   X1_BLTS_PROCS : ALIAS FOR I[3].0;
   XFER1A_BLTS_PRO : ALIAS FOR I[3].6;
   Z200 : MAC_Zone_ML := (ST_xManualModeConditionOK := 1, ST_xZoneError := 1, tmON_480Vca.ACC := 10, tmON_480Vca.EN := 1, tmON_480Vca.DN := 1);
   Z200_ALM : MAC_Zone_ML_ALM := (rgxEmergency[0] := 1, rgxStoppingFault[0] := 63, rgxWarning[0] := 7);
        .rgxEmergency[0].0   // MCC1201.A34KE1.Main Emergency ON
        .rgxStoppingFault[0].0   // Z200.MCC1201.24Vdc Voltage Fault
        .rgxEmergency[0].1   // MCC1201.A33SB1.Main Emergency localization (MCC1201 cabinet)
        .rgxEmergency[0].2   // M203S.A34SB1.Main Emergency localization (operator side)
        .rgxEmergency[0].3   // M203S.A34SB2.Main Emergency localization (far side)
        .rgxStoppingFault[0].1   // Z200.MCC1201.A18QF31/32/33/34.Power supply 24Vdc Fault
        .rgxStoppingFault[0].2   // Z200.MCC1201.A18QF41/42/43/44.Power supply 24Vdc Fault
        .rgxStoppingFault[0].3   // Z200.MCC1201.A19QF11/12/13/14.Power supply 24Vdc Fault
        .rgxStoppingFault[0].4   // Z200.MCC1201.A19QF21/22/23/24.Power supply 24Vdc Fault
        .rgxFault[0].0   // Z200.MCC1201.A155SW1.Ethernet Switch Fault
        .rgxWarning[0].0   // Z200.MCC1201.A11QF1.Power failure 120V Auxiliary
        .rgxWarning[0].1   // Z200.MCC1201.A11QF3.Power failure 120V Auxiliary
        .rgxWarning[0].2   // Z200.MCC1201.A16QF1.Protection power supply conditioner
        .rgxStoppingFault[0].5   // Z200.MCC1201.A18GS1.24Vdc Power Supply Fault
   Z200_HMR : MAC_Zone_ML_HMR := (xZoneAlarm := 1, dZoneState := 1024, dCabinetState := 2, dCleaningState := 2, dManualSpeed_mm_min := 1270);
   Z200_HMW : MAC_Zone_ML_HMW;
   Z200_UPS : ZONE_UPS := (ST_xZoneError := 1, ST_xSelectionManualMode := 1, ST_xConditionOKManualMode := 1, ST_xManualModeAccepted := 1, ST_xZoneEmergency := 1, INPUT_xPowerFailurePLCA := 1, INPUT_xPowerFailurePLCB := 1, AUX_tmOFF_ResetAlarm.PRE := 1000, AUX_tmOFF_ResetAlarm.ACC := 1000, AUX_tmON_24Vdc.PRE := 5000, AUX_tmON_EmergencyOK.PRE := 5000, AUX_tmON_Clutch1feedback.PRE := 1000, AUX_tmON_Clutch2feedback.PRE := 1000); {access None}
   Z200_UPS_ALM : ZONE_UPS_ALM := (rgxEmergency[0] := 1); {access Read Only}
        .rgxEmergency[0].0   // MCC1201.A33KE1.UPS Emergency ON
        .rgxEmergency[0].1   // M203S.A33SB2.UPS Emergency localization (operator side)
        .rgxEmergency[0].2   // M203S.A33SB3.UPS Emergency localization (far side)
        .rgxEmergency[0].3   // M225S.A33SB4.UPS Emergency localization (operator side CS4425)
        .rgxEmergency[0].4   // M225S.A33SB5.UPS Emergency localization (operator side CS4425)
   Z200_UPS_HMR : ZONE_UPS_HMR := (dZoneMode := 1, xZoneAlarm := 1, dZoneState := 1024); {access Read Only}
   Z200_UPS_HMW : ZONE_UPS_HMW;
   Z_ONS_BIT : BOOL[32];   // Temporary Boolean tag created during conversion
END_VAR

PROGRAM _18_STI   (* main routine _18_STI *)

ROUTINE _18_STI   (* ladder *)
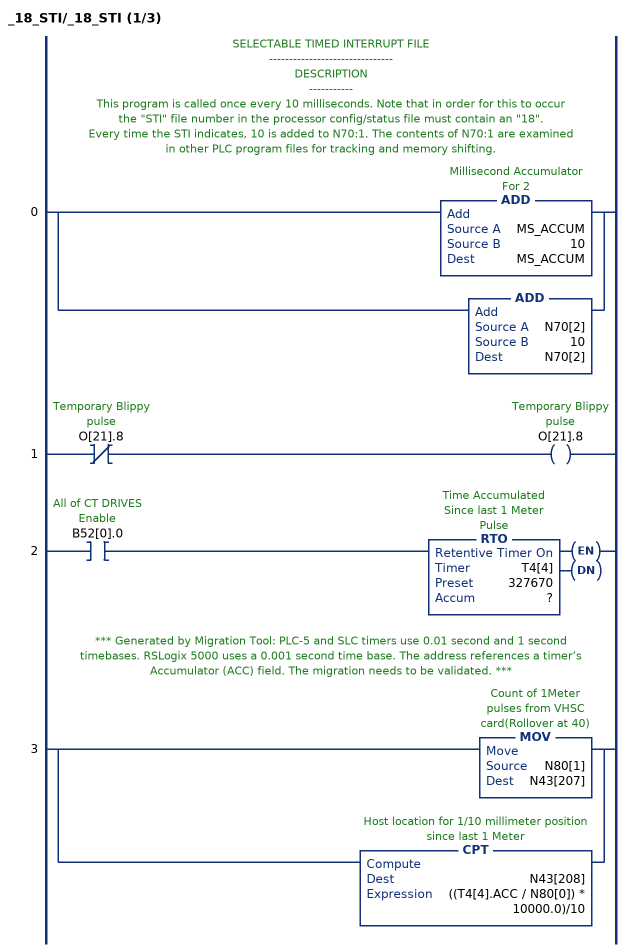
   // SELECTABLE TIMED INTERRUPT FILE
   // -------------------------------
   // DESCRIPTION
   // -----------
   // This program is called once every 10 milliseconds. Note that in order for this to occur
   // the "STI" file number in the processor config/status file must contain an "18".
   // Every time the STI indicates, 10 is added to N70:1. The contents of N70:1 are examined
   // in other PLC program files for tracking and memory shifting.
   0: [ADD(MS_ACCUM,10,MS_ACCUM) ,ADD(N70[2],10,N70[2]) ];
   1: XIO(O[21].8)OTE(O[21].8);
   2: XIC(B52[0].0)RTO(T4[4],?,?);
   // *** Generated by Migration Tool: PLC-5 and SLC timers use 0.01 second and 1 second timebases. RSLogix 5000 uses a 0.001 second time base. The address references a timer’s Accumulator (ACC) field. The migration needs to be validated. ***
   3: [MOV(N80[1],N43[207]) ,CPT(N43[208],((T4[4].ACC / N80[0]) * 10000.0)/10) ];
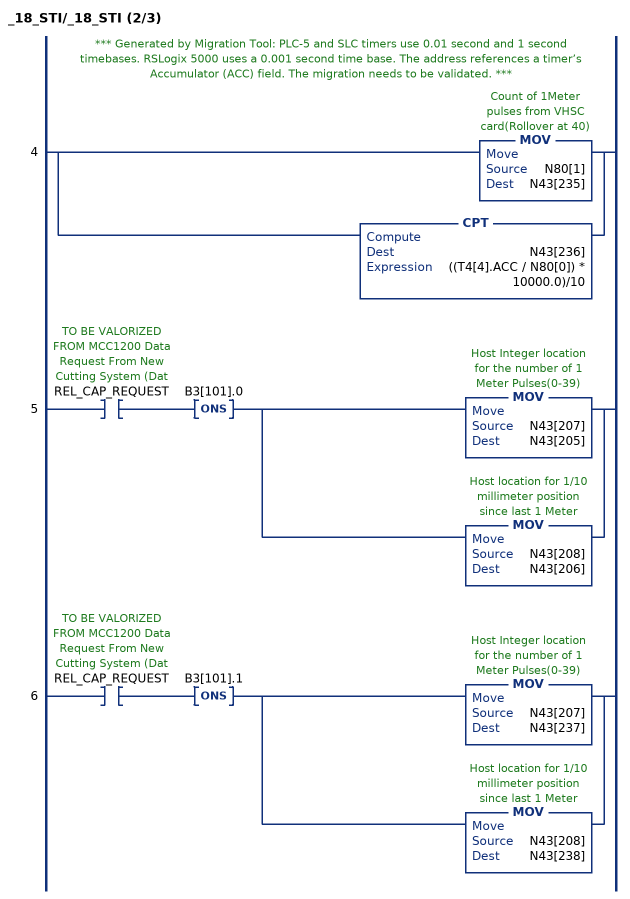
   // *** Generated by Migration Tool: PLC-5 and SLC timers use 0.01 second and 1 second timebases. RSLogix 5000 uses a 0.001 second time base. The address references a timer’s Accumulator (ACC) field. The migration needs to be validated. ***
   4: [MOV(N80[1],N43[235]) ,CPT(N43[236],((T4[4].ACC / N80[0]) * 10000.0)/10) ];
   5: XIC(REL_CAP_REQUEST)ONS(B3[101].0)[MOV(N43[207],N43[205]) ,MOV(N43[208],N43[206]) ];
   6: XIC(REL_CAP_REQUEST)ONS(B3[101].1)[MOV(N43[207],N43[237]) ,MOV(N43[208],N43[238]) ];
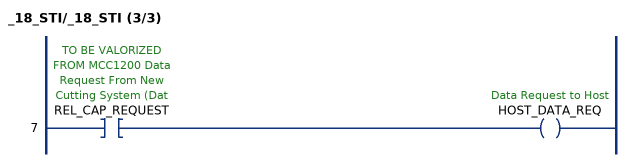
   7: XIC(REL_CAP_REQUEST)OTE(HOST_DATA_REQ);
END_ROUTINE
END_PROGRAM

PROGRAM CommandLogic   (* main routine Main *)
VAR
   TMP_rDummy : REAL;
   TMP_rTarget : REAL;
   TMP_xDummy : BOOL;
   WASHER_ALARM_HORN_RESET : BOOL;
END_VAR

ROUTINE M202_Conveyor_Motion_Output   (* ladder *)
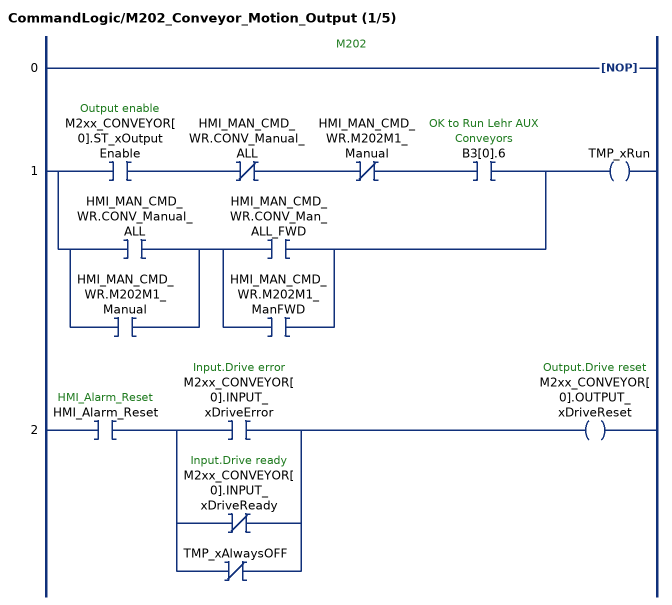
   // M202
   0: NOP();
   1: [XIC(M2xx_CONVEYOR[0].ST_xOutputEnable) XIO(HMI_MAN_CMD_WR.CONV_Manual_ALL) XIO(HMI_MAN_CMD_WR.M202M1_Manual) XIC(B3[0].6) ,[XIC(HMI_MAN_CMD_WR.CONV_Manual_ALL) ,XIC(HMI_MAN_CMD_WR.M202M1_Manual) ] [XIC(HMI_MAN_CMD_WR.CONV_Man_ALL_FWD) ,XIC(HMI_MAN_CMD_WR.M202M1_ManFWD) ] ]OTE(TMP_xRun);
   2: XIC(HMI_Alarm_Reset)[XIC(M2xx_CONVEYOR[0].INPUT_xDriveError) ,XIO(M2xx_CONVEYOR[0].INPUT_xDriveReady) ,XIO(TMP_xAlwaysOFF) ]OTE(M2xx_CONVEYOR[0].OUTPUT_xDriveReset);
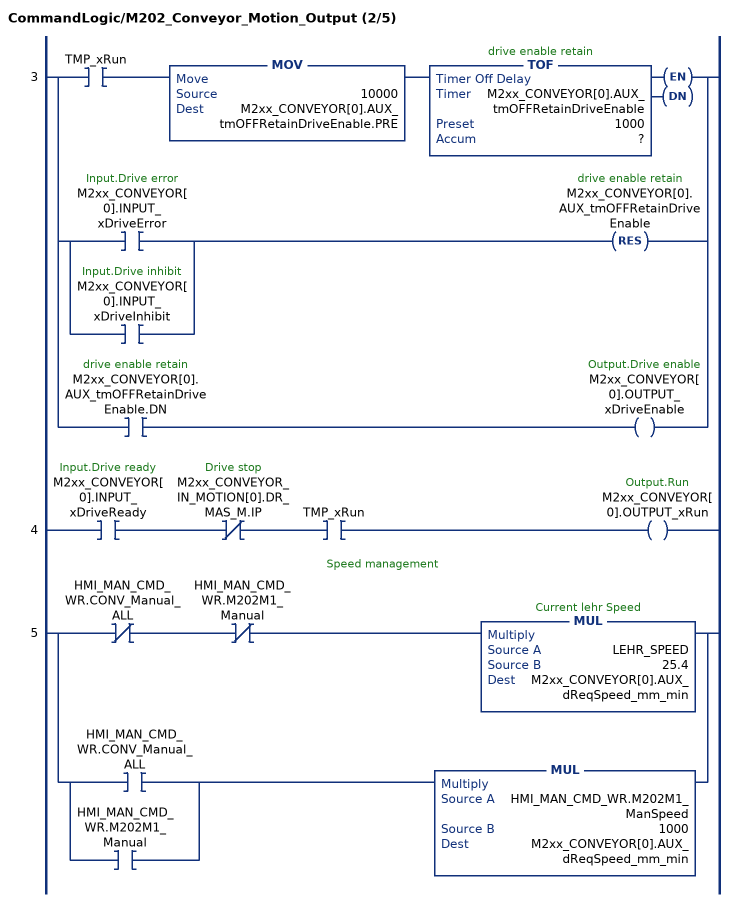
   3: [XIC(TMP_xRun) MOV(10000,M2xx_CONVEYOR[0].AUX_tmOFFRetainDriveEnable.PRE) TOF(M2xx_CONVEYOR[0].AUX_tmOFFRetainDriveEnable,?,?) ,[XIC(M2xx_CONVEYOR[0].INPUT_xDriveError) ,XIC(M2xx_CONVEYOR[0].INPUT_xDriveInhibit) ] RES(M2xx_CONVEYOR[0].AUX_tmOFFRetainDriveEnable) ,XIC(M2xx_CONVEYOR[0].AUX_tmOFFRetainDriveEnable.DN) OTE(M2xx_CONVEYOR[0].OUTPUT_xDriveEnable) ];
   4: XIC(M2xx_CONVEYOR[0].INPUT_xDriveReady)XIO(M2xx_CONVEYOR_IN_MOTION[0].DR_MAS_M.IP)XIC(TMP_xRun)OTE(M2xx_CONVEYOR[0].OUTPUT_xRun);
   // Speed management
   5: [XIO(HMI_MAN_CMD_WR.CONV_Manual_ALL) XIO(HMI_MAN_CMD_WR.M202M1_Manual) MUL(LEHR_SPEED,25.4,M2xx_CONVEYOR[0].AUX_dReqSpeed_mm_min) ,[XIC(HMI_MAN_CMD_WR.CONV_Manual_ALL) ,XIC(HMI_MAN_CMD_WR.M202M1_Manual) ] MUL(HMI_MAN_CMD_WR.M202M1_ManSpeed,1000,M2xx_CONVEYOR[0].AUX_dReqSpeed_mm_min) ];
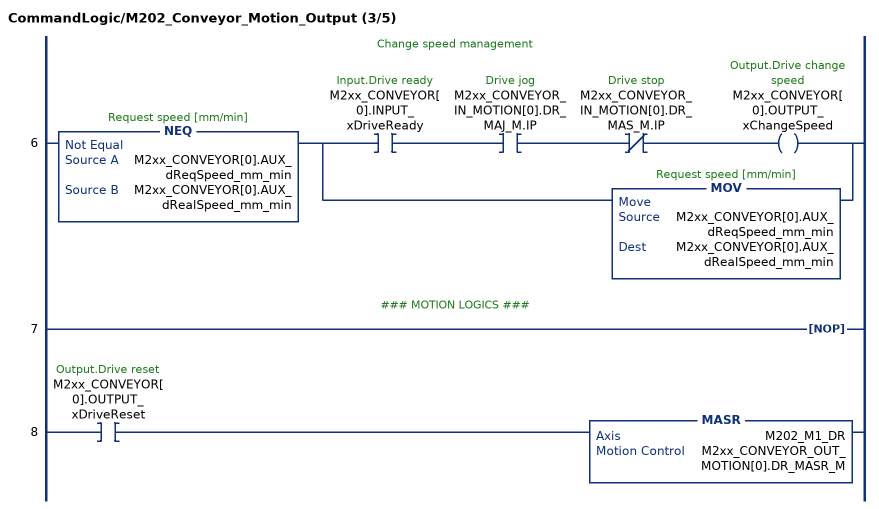
   // Change speed management
   6: NEQ(M2xx_CONVEYOR[0].AUX_dReqSpeed_mm_min,M2xx_CONVEYOR[0].AUX_dRealSpeed_mm_min)[XIC(M2xx_CONVEYOR[0].INPUT_xDriveReady) XIC(M2xx_CONVEYOR_IN_MOTION[0].DR_MAJ_M.IP) XIO(M2xx_CONVEYOR_IN_MOTION[0].DR_MAS_M.IP) OTE(M2xx_CONVEYOR[0].OUTPUT_xChangeSpeed) ,MOV(M2xx_CONVEYOR[0].AUX_dReqSpeed_mm_min,M2xx_CONVEYOR[0].AUX_dRealSpeed_mm_min) ];
   // ### MOTION LOGICS ###
   7: NOP();
   8: XIC(M2xx_CONVEYOR[0].OUTPUT_xDriveReset)MASR(M202_M1_DR,M2xx_CONVEYOR_OUT_MOTION[0].DR_MASR_M);
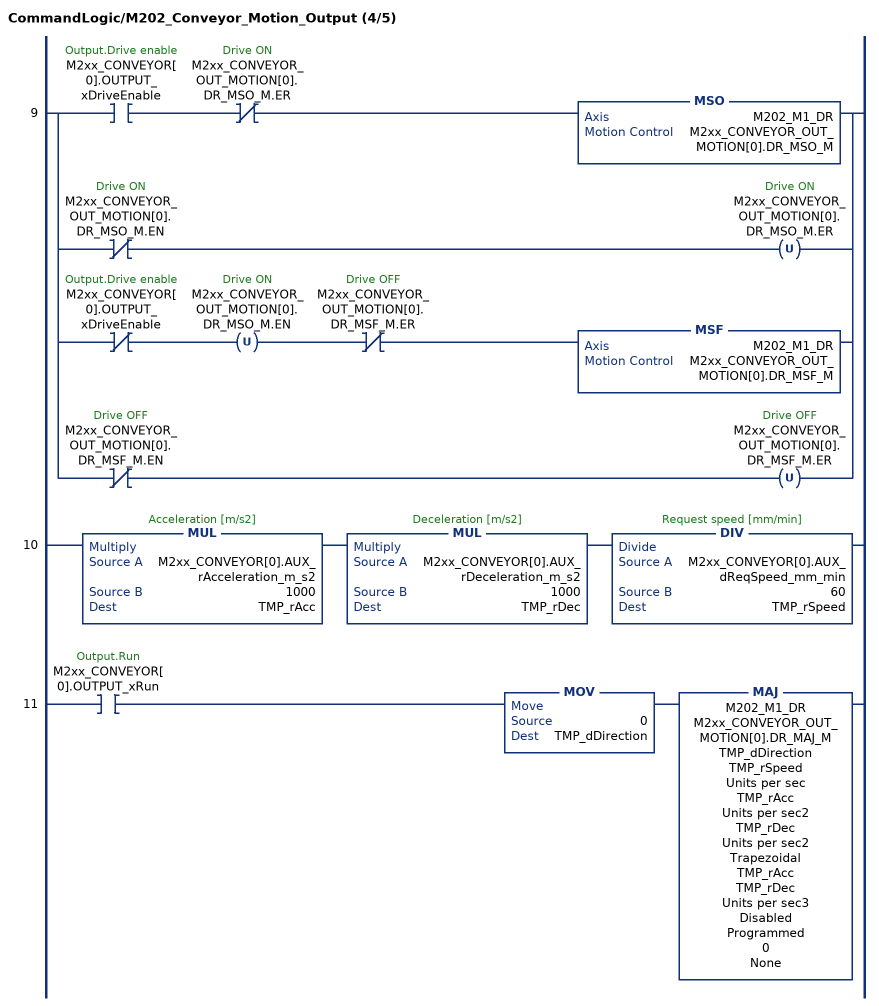
   9: [XIC(M2xx_CONVEYOR[0].OUTPUT_xDriveEnable) XIO(M2xx_CONVEYOR_OUT_MOTION[0].DR_MSO_M.ER) MSO(M202_M1_DR,M2xx_CONVEYOR_OUT_MOTION[0].DR_MSO_M) ,XIO(M2xx_CONVEYOR_OUT_MOTION[0].DR_MSO_M.EN) OTU(M2xx_CONVEYOR_OUT_MOTION[0].DR_MSO_M.ER) ,XIO(M2xx_CONVEYOR[0].OUTPUT_xDriveEnable) OTU(M2xx_CONVEYOR_OUT_MOTION[0].DR_MSO_M.EN) XIO(M2xx_CONVEYOR_OUT_MOTION[0].DR_MSF_M.ER) MSF(M202_M1_DR,M2xx_CONVEYOR_OUT_MOTION[0].DR_MSF_M) ,XIO(M2xx_CONVEYOR_OUT_MOTION[0].DR_MSF_M.EN) OTU(M2xx_CONVEYOR_OUT_MOTION[0].DR_MSF_M.ER) ];
   10: MUL(M2xx_CONVEYOR[0].AUX_rAcceleration_m_s2,1000,TMP_rAcc)MUL(M2xx_CONVEYOR[0].AUX_rDeceleration_m_s2,1000,TMP_rDec)DIV(M2xx_CONVEYOR[0].AUX_dReqSpeed_mm_min,60,TMP_rSpeed);
   11: XIC(M2xx_CONVEYOR[0].OUTPUT_xRun)MOV(0,TMP_dDirection)MAJ(M202_M1_DR,M2xx_CONVEYOR_OUT_MOTION[0].DR_MAJ_M,TMP_dDirection,TMP_rSpeed,Units per sec,TMP_rAcc,Units per sec2,TMP_rDec,Units per sec2,Trapezoidal,TMP_rAcc,TMP_rDec,Units per sec3,Disabled,Programmed,0,None);
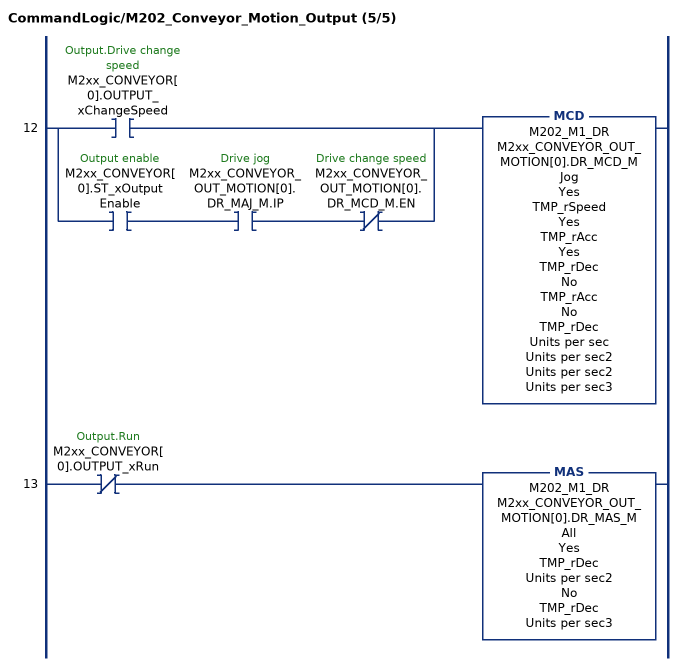
   12: [XIC(M2xx_CONVEYOR[0].OUTPUT_xChangeSpeed) ,XIC(M2xx_CONVEYOR[0].ST_xOutputEnable) XIC(M2xx_CONVEYOR_OUT_MOTION[0].DR_MAJ_M.IP) XIO(M2xx_CONVEYOR_OUT_MOTION[0].DR_MCD_M.EN) ]MCD(M202_M1_DR,M2xx_CONVEYOR_OUT_MOTION[0].DR_MCD_M,Jog,Yes,TMP_rSpeed,Yes,TMP_rAcc,Yes,TMP_rDec,No,TMP_rAcc,No,TMP_rDec,Units per sec,Units per sec2,Units per sec2,Units per sec3);
   13: XIO(M2xx_CONVEYOR[0].OUTPUT_xRun)MAS(M202_M1_DR,M2xx_CONVEYOR_OUT_MOTION[0].DR_MAS_M,All,Yes,TMP_rDec,Units per sec2,No,TMP_rDec,Units per sec3);
END_ROUTINE

ROUTINE M203_Conveyor_Motion_Output   (* ladder *)
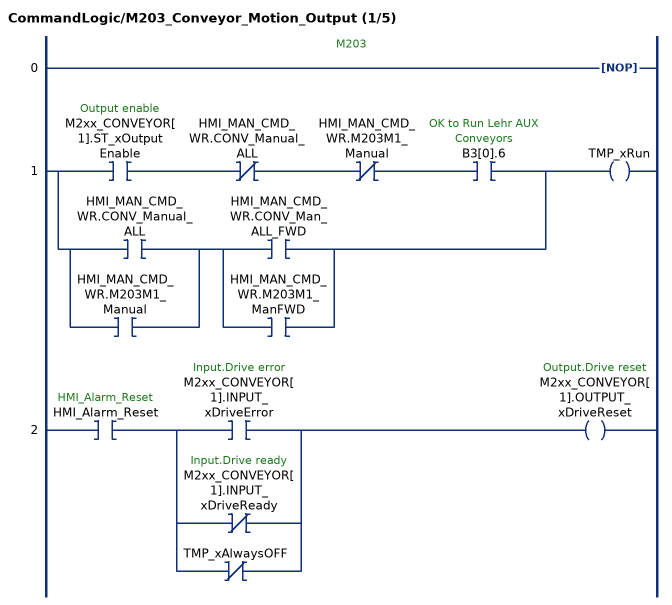
   // M203
   0: NOP();
   1: [XIC(M2xx_CONVEYOR[1].ST_xOutputEnable) XIO(HMI_MAN_CMD_WR.CONV_Manual_ALL) XIO(HMI_MAN_CMD_WR.M203M1_Manual) XIC(B3[0].6) ,[XIC(HMI_MAN_CMD_WR.CONV_Manual_ALL) ,XIC(HMI_MAN_CMD_WR.M203M1_Manual) ] [XIC(HMI_MAN_CMD_WR.CONV_Man_ALL_FWD) ,XIC(HMI_MAN_CMD_WR.M203M1_ManFWD) ] ]OTE(TMP_xRun);
   2: XIC(HMI_Alarm_Reset)[XIC(M2xx_CONVEYOR[1].INPUT_xDriveError) ,XIO(M2xx_CONVEYOR[1].INPUT_xDriveReady) ,XIO(TMP_xAlwaysOFF) ]OTE(M2xx_CONVEYOR[1].OUTPUT_xDriveReset);
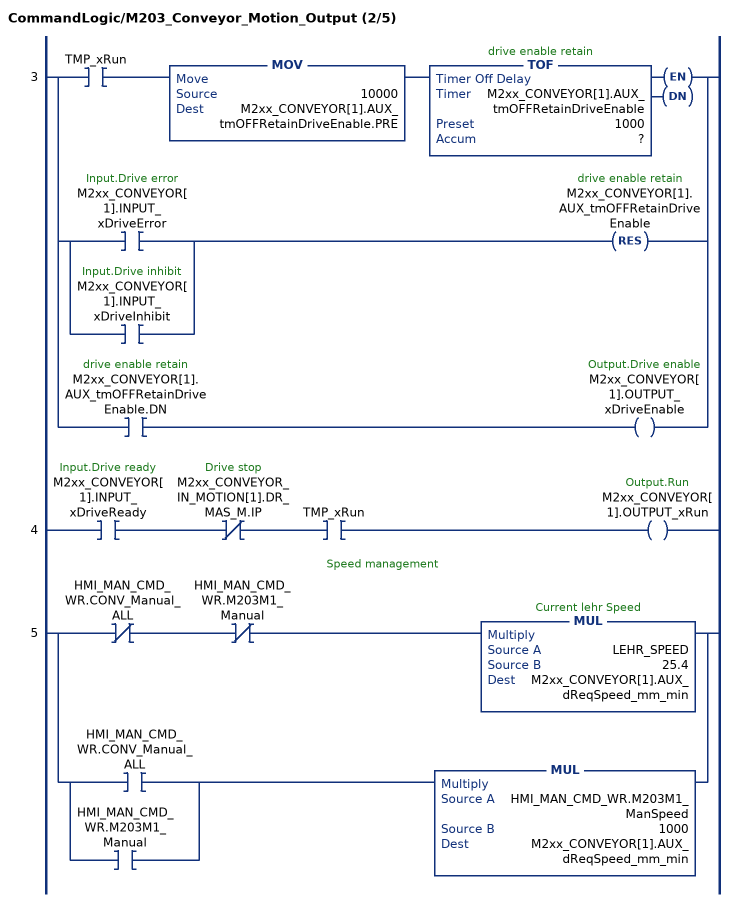
   3: [XIC(TMP_xRun) MOV(10000,M2xx_CONVEYOR[1].AUX_tmOFFRetainDriveEnable.PRE) TOF(M2xx_CONVEYOR[1].AUX_tmOFFRetainDriveEnable,?,?) ,[XIC(M2xx_CONVEYOR[1].INPUT_xDriveError) ,XIC(M2xx_CONVEYOR[1].INPUT_xDriveInhibit) ] RES(M2xx_CONVEYOR[1].AUX_tmOFFRetainDriveEnable) ,XIC(M2xx_CONVEYOR[1].AUX_tmOFFRetainDriveEnable.DN) OTE(M2xx_CONVEYOR[1].OUTPUT_xDriveEnable) ];
   4: XIC(M2xx_CONVEYOR[1].INPUT_xDriveReady)XIO(M2xx_CONVEYOR_IN_MOTION[1].DR_MAS_M.IP)XIC(TMP_xRun)OTE(M2xx_CONVEYOR[1].OUTPUT_xRun);
   // Speed management
   5: [XIO(HMI_MAN_CMD_WR.CONV_Manual_ALL) XIO(HMI_MAN_CMD_WR.M203M1_Manual) MUL(LEHR_SPEED,25.4,M2xx_CONVEYOR[1].AUX_dReqSpeed_mm_min) ,[XIC(HMI_MAN_CMD_WR.CONV_Manual_ALL) ,XIC(HMI_MAN_CMD_WR.M203M1_Manual) ] MUL(HMI_MAN_CMD_WR.M203M1_ManSpeed,1000,M2xx_CONVEYOR[1].AUX_dReqSpeed_mm_min) ];
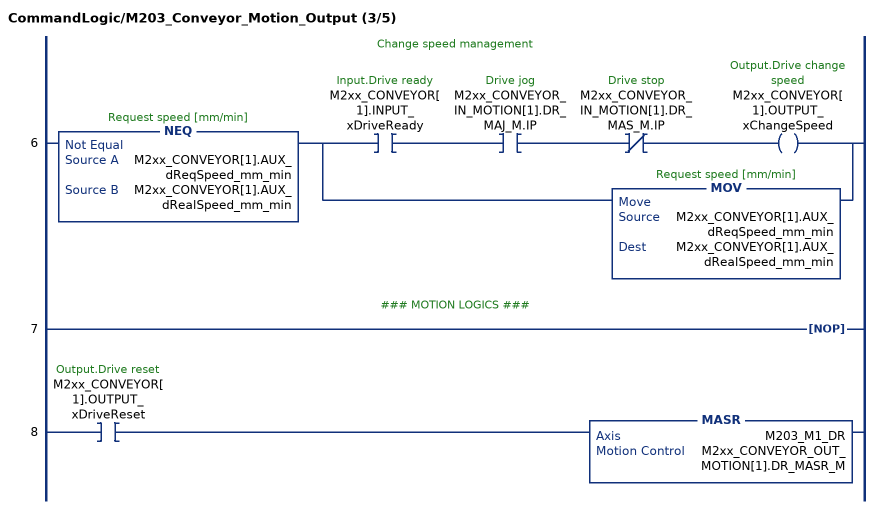
   // Change speed management
   6: NEQ(M2xx_CONVEYOR[1].AUX_dReqSpeed_mm_min,M2xx_CONVEYOR[1].AUX_dRealSpeed_mm_min)[XIC(M2xx_CONVEYOR[1].INPUT_xDriveReady) XIC(M2xx_CONVEYOR_IN_MOTION[1].DR_MAJ_M.IP) XIO(M2xx_CONVEYOR_IN_MOTION[1].DR_MAS_M.IP) OTE(M2xx_CONVEYOR[1].OUTPUT_xChangeSpeed) ,MOV(M2xx_CONVEYOR[1].AUX_dReqSpeed_mm_min,M2xx_CONVEYOR[1].AUX_dRealSpeed_mm_min) ];
   // ### MOTION LOGICS ###
   7: NOP();
   8: XIC(M2xx_CONVEYOR[1].OUTPUT_xDriveReset)MASR(M203_M1_DR,M2xx_CONVEYOR_OUT_MOTION[1].DR_MASR_M);
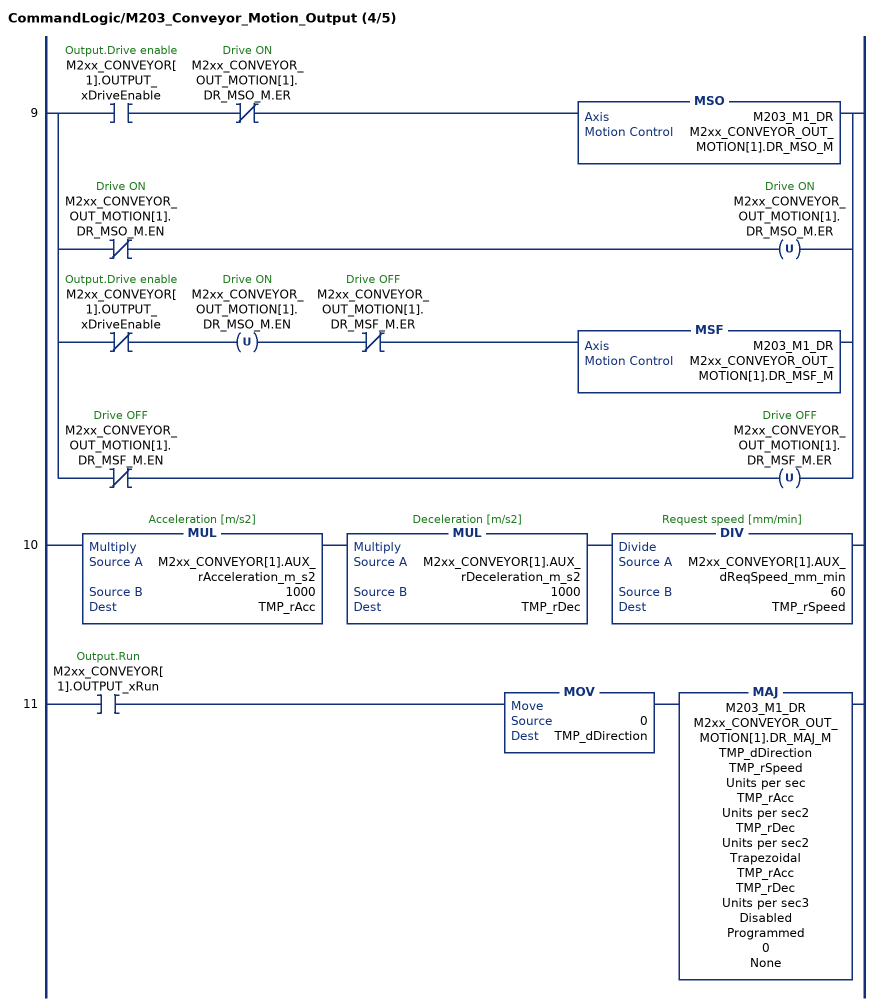
   9: [XIC(M2xx_CONVEYOR[1].OUTPUT_xDriveEnable) XIO(M2xx_CONVEYOR_OUT_MOTION[1].DR_MSO_M.ER) MSO(M203_M1_DR,M2xx_CONVEYOR_OUT_MOTION[1].DR_MSO_M) ,XIO(M2xx_CONVEYOR_OUT_MOTION[1].DR_MSO_M.EN) OTU(M2xx_CONVEYOR_OUT_MOTION[1].DR_MSO_M.ER) ,XIO(M2xx_CONVEYOR[1].OUTPUT_xDriveEnable) OTU(M2xx_CONVEYOR_OUT_MOTION[1].DR_MSO_M.EN) XIO(M2xx_CONVEYOR_OUT_MOTION[1].DR_MSF_M.ER) MSF(M203_M1_DR,M2xx_CONVEYOR_OUT_MOTION[1].DR_MSF_M) ,XIO(M2xx_CONVEYOR_OUT_MOTION[1].DR_MSF_M.EN) OTU(M2xx_CONVEYOR_OUT_MOTION[1].DR_MSF_M.ER) ];
   10: MUL(M2xx_CONVEYOR[1].AUX_rAcceleration_m_s2,1000,TMP_rAcc)MUL(M2xx_CONVEYOR[1].AUX_rDeceleration_m_s2,1000,TMP_rDec)DIV(M2xx_CONVEYOR[1].AUX_dReqSpeed_mm_min,60,TMP_rSpeed);
   11: XIC(M2xx_CONVEYOR[1].OUTPUT_xRun)MOV(0,TMP_dDirection)MAJ(M203_M1_DR,M2xx_CONVEYOR_OUT_MOTION[1].DR_MAJ_M,TMP_dDirection,TMP_rSpeed,Units per sec,TMP_rAcc,Units per sec2,TMP_rDec,Units per sec2,Trapezoidal,TMP_rAcc,TMP_rDec,Units per sec3,Disabled,Programmed,0,None);
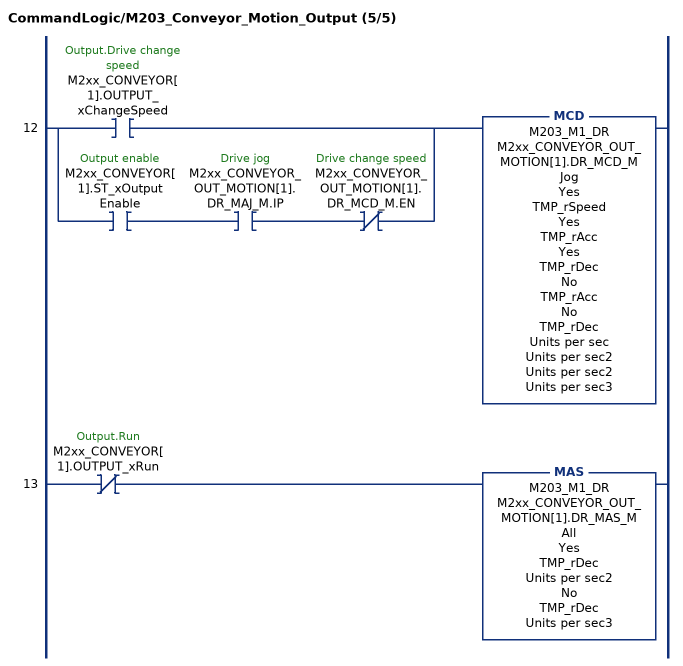
   12: [XIC(M2xx_CONVEYOR[1].OUTPUT_xChangeSpeed) ,XIC(M2xx_CONVEYOR[1].ST_xOutputEnable) XIC(M2xx_CONVEYOR_OUT_MOTION[1].DR_MAJ_M.IP) XIO(M2xx_CONVEYOR_OUT_MOTION[1].DR_MCD_M.EN) ]MCD(M203_M1_DR,M2xx_CONVEYOR_OUT_MOTION[1].DR_MCD_M,Jog,Yes,TMP_rSpeed,Yes,TMP_rAcc,Yes,TMP_rDec,No,TMP_rAcc,No,TMP_rDec,Units per sec,Units per sec2,Units per sec2,Units per sec3);
   13: XIO(M2xx_CONVEYOR[1].OUTPUT_xRun)MAS(M203_M1_DR,M2xx_CONVEYOR_OUT_MOTION[1].DR_MAS_M,All,Yes,TMP_rDec,Units per sec2,No,TMP_rDec,Units per sec3);
END_ROUTINE

ROUTINE M203_DropConveyor_Output   (* ladder *)
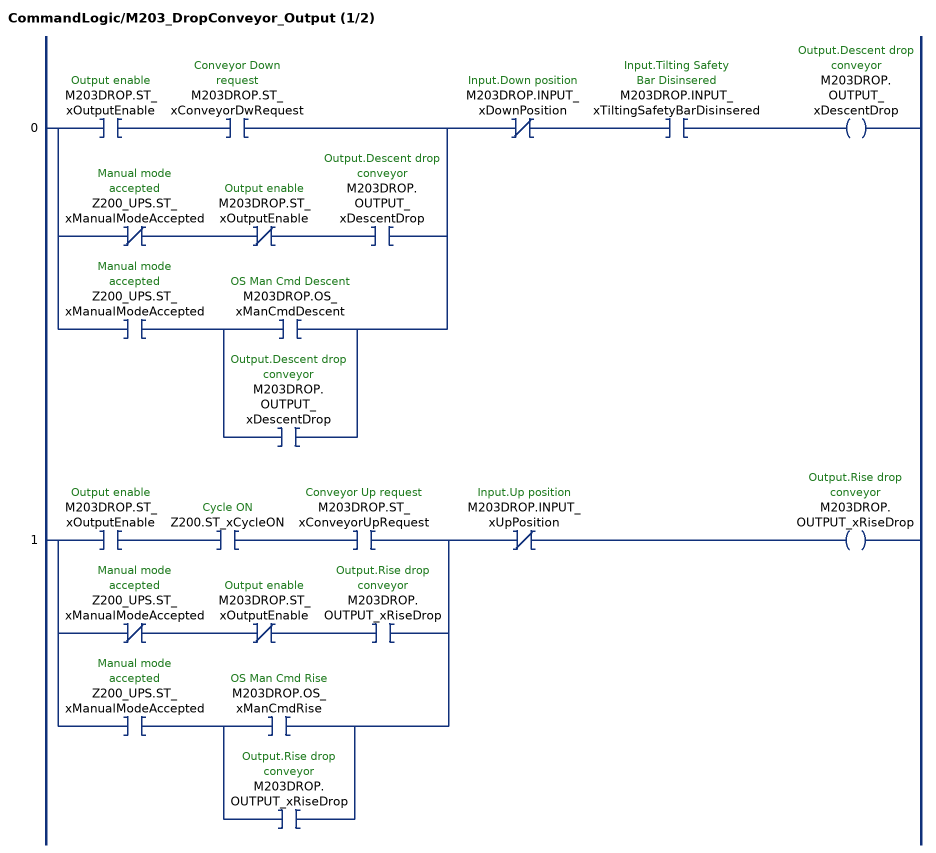
   0: [XIC(M203DROP.ST_xOutputEnable) XIC(M203DROP.ST_xConveyorDwRequest) ,XIO(Z200_UPS.ST_xManualModeAccepted) XIO(M203DROP.ST_xOutputEnable) XIC(M203DROP.OUTPUT_xDescentDrop) ,XIC(Z200_UPS.ST_xManualModeAccepted) [XIC(M203DROP.OS_xManCmdDescent) ,XIC(M203DROP.OUTPUT_xDescentDrop) ] ]XIO(M203DROP.INPUT_xDownPosition)XIC(M203DROP.INPUT_xTiltingSafetyBarDisinsered)OTE(M203DROP.OUTPUT_xDescentDrop);
   1: [XIC(M203DROP.ST_xOutputEnable) XIC(Z200.ST_xCycleON) XIC(M203DROP.ST_xConveyorUpRequest) ,XIO(Z200_UPS.ST_xManualModeAccepted) XIO(M203DROP.ST_xOutputEnable) XIC(M203DROP.OUTPUT_xRiseDrop) ,XIC(Z200_UPS.ST_xManualModeAccepted) [XIC(M203DROP.OS_xManCmdRise) ,XIC(M203DROP.OUTPUT_xRiseDrop) ] ]XIO(M203DROP.INPUT_xUpPosition)OTE(M203DROP.OUTPUT_xRiseDrop);
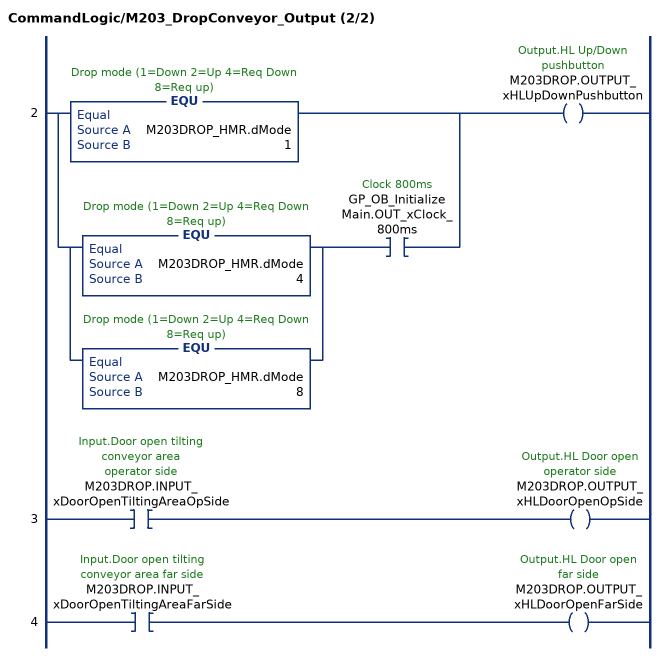
   2: [EQU(M203DROP_HMR.dMode,1) ,[EQU(M203DROP_HMR.dMode,4) ,EQU(M203DROP_HMR.dMode,8) ] XIC(GP_OB_InitializeMain.OUT_xClock_800ms) ]OTE(M203DROP.OUTPUT_xHLUpDownPushbutton);
   3: XIC(M203DROP.INPUT_xDoorOpenTiltingAreaOpSide)OTE(M203DROP.OUTPUT_xHLDoorOpenOpSide);
   4: XIC(M203DROP.INPUT_xDoorOpenTiltingAreaFarSide)OTE(M203DROP.OUTPUT_xHLDoorOpenFarSide);
END_ROUTINE

ROUTINE M204_Conveyor_Motion_Output   (* ladder *)
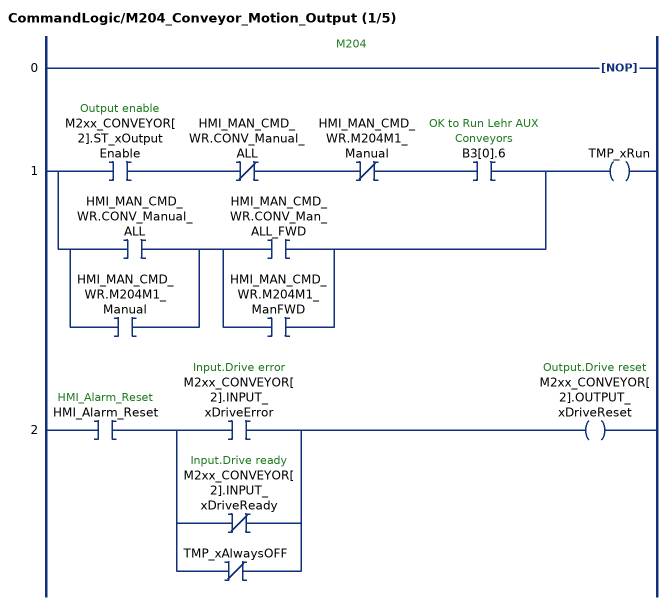
   // M204
   0: NOP();
   1: [XIC(M2xx_CONVEYOR[2].ST_xOutputEnable) XIO(HMI_MAN_CMD_WR.CONV_Manual_ALL) XIO(HMI_MAN_CMD_WR.M204M1_Manual) XIC(B3[0].6) ,[XIC(HMI_MAN_CMD_WR.CONV_Manual_ALL) ,XIC(HMI_MAN_CMD_WR.M204M1_Manual) ] [XIC(HMI_MAN_CMD_WR.CONV_Man_ALL_FWD) ,XIC(HMI_MAN_CMD_WR.M204M1_ManFWD) ] ]OTE(TMP_xRun);
   2: XIC(HMI_Alarm_Reset)[XIC(M2xx_CONVEYOR[2].INPUT_xDriveError) ,XIO(M2xx_CONVEYOR[2].INPUT_xDriveReady) ,XIO(TMP_xAlwaysOFF) ]OTE(M2xx_CONVEYOR[2].OUTPUT_xDriveReset);
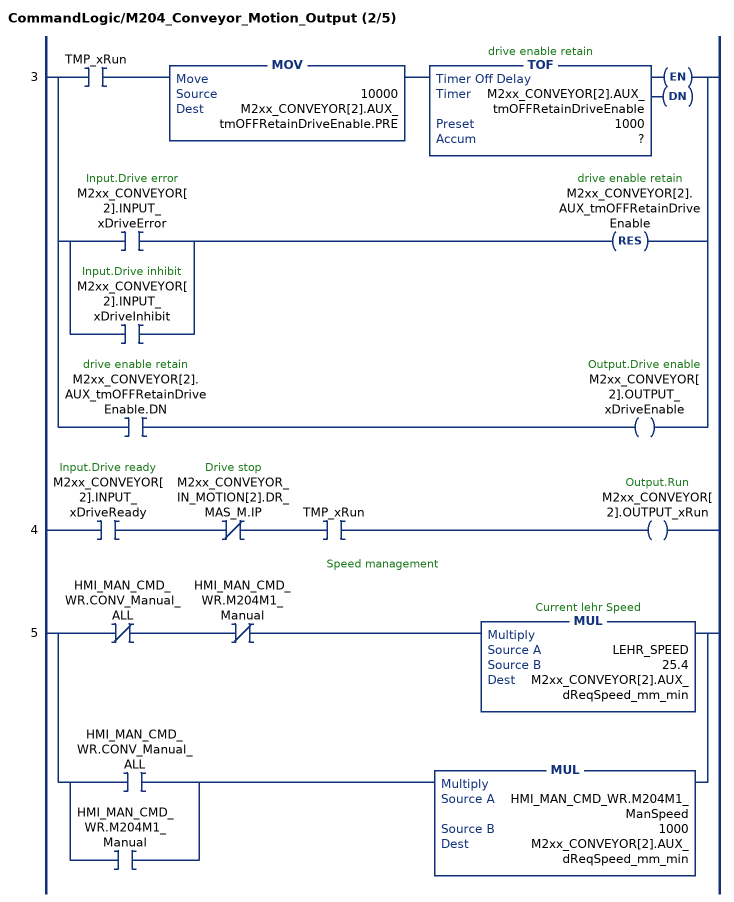
   3: [XIC(TMP_xRun) MOV(10000,M2xx_CONVEYOR[2].AUX_tmOFFRetainDriveEnable.PRE) TOF(M2xx_CONVEYOR[2].AUX_tmOFFRetainDriveEnable,?,?) ,[XIC(M2xx_CONVEYOR[2].INPUT_xDriveError) ,XIC(M2xx_CONVEYOR[2].INPUT_xDriveInhibit) ] RES(M2xx_CONVEYOR[2].AUX_tmOFFRetainDriveEnable) ,XIC(M2xx_CONVEYOR[2].AUX_tmOFFRetainDriveEnable.DN) OTE(M2xx_CONVEYOR[2].OUTPUT_xDriveEnable) ];
   4: XIC(M2xx_CONVEYOR[2].INPUT_xDriveReady)XIO(M2xx_CONVEYOR_IN_MOTION[2].DR_MAS_M.IP)XIC(TMP_xRun)OTE(M2xx_CONVEYOR[2].OUTPUT_xRun);
   // Speed management
   5: [XIO(HMI_MAN_CMD_WR.CONV_Manual_ALL) XIO(HMI_MAN_CMD_WR.M204M1_Manual) MUL(LEHR_SPEED,25.4,M2xx_CONVEYOR[2].AUX_dReqSpeed_mm_min) ,[XIC(HMI_MAN_CMD_WR.CONV_Manual_ALL) ,XIC(HMI_MAN_CMD_WR.M204M1_Manual) ] MUL(HMI_MAN_CMD_WR.M204M1_ManSpeed,1000,M2xx_CONVEYOR[2].AUX_dReqSpeed_mm_min) ];
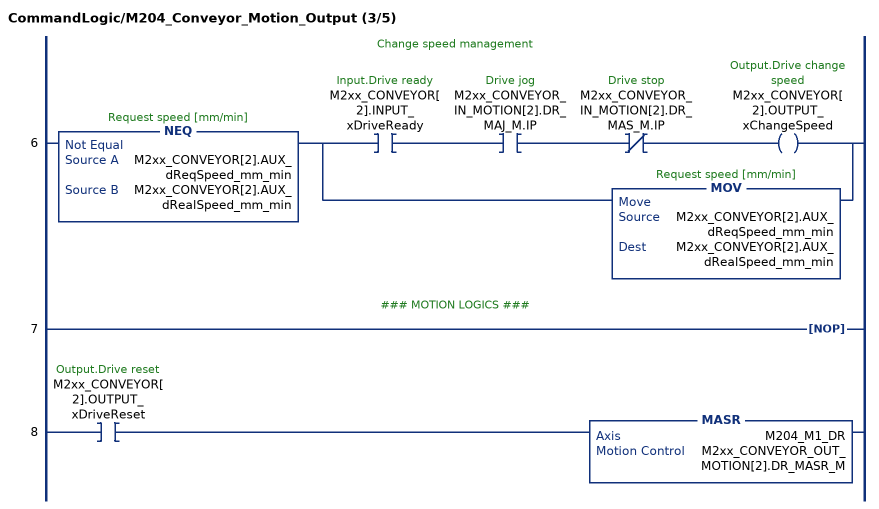
   // Change speed management
   6: NEQ(M2xx_CONVEYOR[2].AUX_dReqSpeed_mm_min,M2xx_CONVEYOR[2].AUX_dRealSpeed_mm_min)[XIC(M2xx_CONVEYOR[2].INPUT_xDriveReady) XIC(M2xx_CONVEYOR_IN_MOTION[2].DR_MAJ_M.IP) XIO(M2xx_CONVEYOR_IN_MOTION[2].DR_MAS_M.IP) OTE(M2xx_CONVEYOR[2].OUTPUT_xChangeSpeed) ,MOV(M2xx_CONVEYOR[2].AUX_dReqSpeed_mm_min,M2xx_CONVEYOR[2].AUX_dRealSpeed_mm_min) ];
   // ### MOTION LOGICS ###
   7: NOP();
   8: XIC(M2xx_CONVEYOR[2].OUTPUT_xDriveReset)MASR(M204_M1_DR,M2xx_CONVEYOR_OUT_MOTION[2].DR_MASR_M);
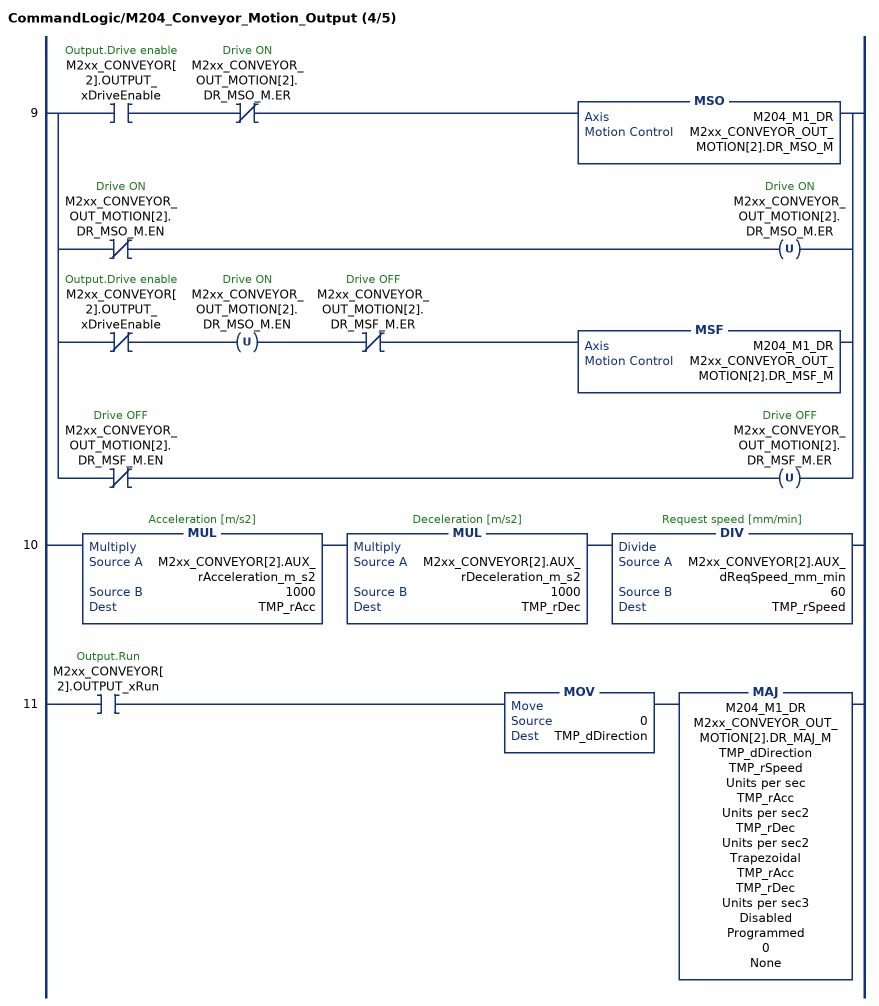
   9: [XIC(M2xx_CONVEYOR[2].OUTPUT_xDriveEnable) XIO(M2xx_CONVEYOR_OUT_MOTION[2].DR_MSO_M.ER) MSO(M204_M1_DR,M2xx_CONVEYOR_OUT_MOTION[2].DR_MSO_M) ,XIO(M2xx_CONVEYOR_OUT_MOTION[2].DR_MSO_M.EN) OTU(M2xx_CONVEYOR_OUT_MOTION[2].DR_MSO_M.ER) ,XIO(M2xx_CONVEYOR[2].OUTPUT_xDriveEnable) OTU(M2xx_CONVEYOR_OUT_MOTION[2].DR_MSO_M.EN) XIO(M2xx_CONVEYOR_OUT_MOTION[2].DR_MSF_M.ER) MSF(M204_M1_DR,M2xx_CONVEYOR_OUT_MOTION[2].DR_MSF_M) ,XIO(M2xx_CONVEYOR_OUT_MOTION[2].DR_MSF_M.EN) OTU(M2xx_CONVEYOR_OUT_MOTION[2].DR_MSF_M.ER) ];
   10: MUL(M2xx_CONVEYOR[2].AUX_rAcceleration_m_s2,1000,TMP_rAcc)MUL(M2xx_CONVEYOR[2].AUX_rDeceleration_m_s2,1000,TMP_rDec)DIV(M2xx_CONVEYOR[2].AUX_dReqSpeed_mm_min,60,TMP_rSpeed);
   11: XIC(M2xx_CONVEYOR[2].OUTPUT_xRun)MOV(0,TMP_dDirection)MAJ(M204_M1_DR,M2xx_CONVEYOR_OUT_MOTION[2].DR_MAJ_M,TMP_dDirection,TMP_rSpeed,Units per sec,TMP_rAcc,Units per sec2,TMP_rDec,Units per sec2,Trapezoidal,TMP_rAcc,TMP_rDec,Units per sec3,Disabled,Programmed,0,None);
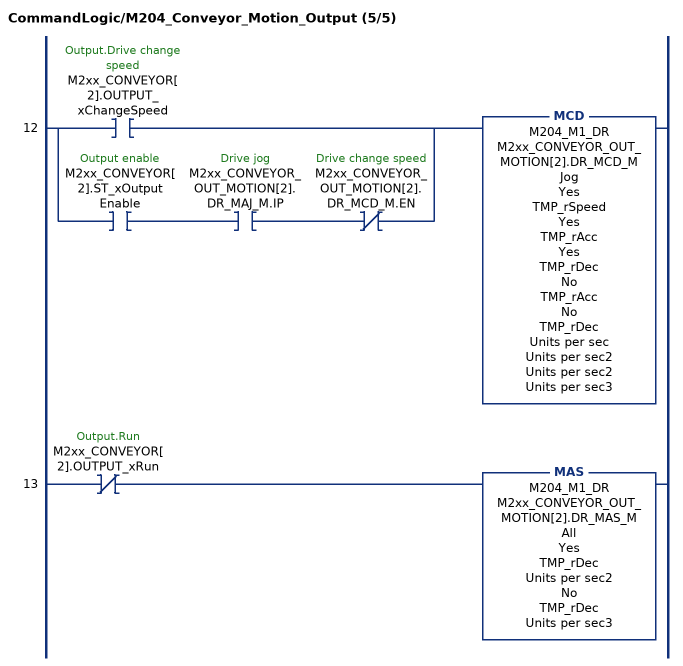
   12: [XIC(M2xx_CONVEYOR[2].OUTPUT_xChangeSpeed) ,XIC(M2xx_CONVEYOR[2].ST_xOutputEnable) XIC(M2xx_CONVEYOR_OUT_MOTION[2].DR_MAJ_M.IP) XIO(M2xx_CONVEYOR_OUT_MOTION[2].DR_MCD_M.EN) ]MCD(M204_M1_DR,M2xx_CONVEYOR_OUT_MOTION[2].DR_MCD_M,Jog,Yes,TMP_rSpeed,Yes,TMP_rAcc,Yes,TMP_rDec,No,TMP_rAcc,No,TMP_rDec,Units per sec,Units per sec2,Units per sec2,Units per sec3);
   13: XIO(M2xx_CONVEYOR[2].OUTPUT_xRun)MAS(M204_M1_DR,M2xx_CONVEYOR_OUT_MOTION[2].DR_MAS_M,All,Yes,TMP_rDec,Units per sec2,No,TMP_rDec,Units per sec3);
END_ROUTINE
